(* Logix 5000 project; controller PLC_MCC1300_75F1 vendor 1 type 14 code 166 rev 32.11; software revision 32.04; part 66 of 83 *)
(* tags used below, declared in another part *)
   CM_ConveyorStackerToLine_JS1_Sync : CM_ConveyorStackerToLine;
   GP_AccessArea_M316S_STC : GP_AccessArea_STC;
   GP_ScadaPlate : GP_ScadaPlate;
   Gp_SpaceConvUtilities_V1 : GP_SpaceConvUtilities_V1;
   M310B : MAC_Conveyor;
   M312 : MAC_Conveyor_Single;
   M312_Data : UDT_Convoy_SL;
   M315A_SpaceConv_Utilities : SpaceConv_Utilities;
   M316 : MAC_Conveyor;
   M316_ALM : MAC_Conveyor_ALM;
   M316_Data : UDT_Convoy_SL;
   M316_HMR : MAC_Conveyor_HMR;
   M316_HMW : MAC_Conveyor_HMW;
   M316_M1_DR : AXIS_CIP_DRIVE;
   M316_SpaceConv_Utilities : SpaceConv_Utilities;
   M316_TON_Synchro_timeout : TIMER;
   M316_xSendCulletReqActive : BOOL;
   M316_xSensorTimeout : BOOL;
   M316A : MAC_Rotator;
   M316A_ALM : MAC_Rotator_ALM;
   M316A_Data : UDT_Convoy_SL;
   M316A_M1_DR_IN_MAM : MOTION_INSTRUCTION;
   M316A_TmON1 : TIMER;
   M316M317_OffsetBaricentre_cmm : DINT;
   M317 : MAC_Conveyor_Single;
   M317_ALM : MAC_Conveyor_ALM;
   M317_Data : UDT_Convoy_SL;
   M317_M2_DR_OUT_MAM : MOTION_INSTRUCTION;
   M317_M3_DR_OUT_MAM : MOTION_INSTRUCTION;
   M317_SpaceConv_Utilities : SpaceConv_Utilities;
   O : INT[128];
   TMP_d : DINT;
   TMP_SendToCullet : BOOL;
   TMP_xConveyorOfStartCleaning : BOOL;
   TMP_xEnableZoneCleaning : BOOL;
   TMP_xLiteThisDestPresent : BOOL;
   xAlwaysOFF : BOOL;
   xAlwaysON : BOOL;
   Z402 : MAC_Zone;
   Z402_HMI_rgtPlateScada_Internal : HMI_LiteData[5,2,7];
   Z402S_INPUT_xSafetyAreaPopup : BOOL;
   Z402S_INPUT_xSafetyAreaRotator : BOOL;
(* MainProgram, continued *)

   // Phase in progress
   48: NEQ(M316.PH_x,0)OTE(M316.ST_xPhasesInProgress);
   // #####_CLEANING_#####
   49: NOP();
   // Cleaning Reset
   50: XIC(M316.ST_xCleaningAccepted)[XIC(Z402.ST_xCleaningAccepted) ,XIO(TMP_xConveyorOfStartCleaning) ][XIC(M316.ST_xIdPlatePresence) OTL(TMP_SendToCullet) FLL(0,M316_Data,1) FLL(0,M316A_Data,1) ,MOV(0,M316A.PH_x) MOV(0,M316.PH_x) OTU(M316.ST_xPlatePresence) ];
   // Redestination lites
   // -
   // -
   51: [XIO(M316.ST_xPhasesInProgress) XIC(M312.ST_xAux1) ,XIC(M316_xSendCulletReqActive) [XIC(xAlwaysOFF) XIC(M316.PH_x.0) ,XIC(xAlwaysOFF) XIC(M316.PH_x.1) ,XIO(M316.ST_xPhasesInProgress) ] ]XIC(TMP_xLiteThisDestPresent)OTL(TMP_SendToCullet);
   // Initial condition OK
   52: XIC(Z402.ST_xConditionOkPhaseAdvancement)XIC(M316.ST_xOutputEnable)XIO(M316_HMW.xEnableDisableManualCommand)XIO(M316.ST_xReqCleaning)XIO(M316.ST_xCleaningAccepted)XIO(M316.ST_xStopNextCycleFault)XIO(M316.ST_xVirtualDoorEnabled)XIO(M316.PH_x.0)[XIO(M316.ST_xPhasesInProgress) XIO(M316.ST_xPlatePresence) XIO(M316.ST_xIdPlatePresence) XIC(M316A.INPUT_xLowPosition) ,XIC(M316.ST_xCycleLoadUnload) XIC(M316.PH_x.8) XIC(M316.OUTPUT_xRun_M1) GRT(M316_SpaceConv_Utilities.O_dTailPosition_cmm,M316_SpaceConv_Utilities.O_dPresetLoadUnload_cmm) GRT(M316_SpaceConv_Utilities.O_dTailPosition_cmm,380000) XIO(M316.ST_xIdPlatePresence) XIO(M312.INPUT_xSyncroPhotocell_1) ]XIO(CM_ConveyorStackerToLine_JS1_Sync.xRequestReturnInLine)XIO(GP_AccessArea_M316S_STC.ST_xAccessRequest)XIO(GP_AccessArea_M316S_STC.ST_xAccessAccepted)OTE(M316.ST_xInitialConditionOK);
   // #### Plate reentry ####
   53: NOP();
   // Initial condition reentry
   54: XIC(Z402.ST_xConditionOkPhaseAdvancement)XIC(M316.ST_xOutputEnable)XIO(M316_HMW.xEnableDisableManualCommand)XIO(M316.ST_xReqCleaning)XIO(M316.ST_xCleaningAccepted)XIO(M316.ST_xStopNextCycleFault)XIO(M312.ST_xVirtualDoorEnabled)XIO(M316.ST_xPhasesInProgress)XIO(M316.ST_xPlatePresence)XIO(M316.ST_xIdPlatePresence)XIC(M316A.INPUT_xLowPosition)XIO(GP_AccessArea_M316S_STC.ST_xAccessRequest)XIO(GP_AccessArea_M316S_STC.ST_xAccessAccepted)XIC(Z402S_INPUT_xSafetyAreaPopup)OTE(M316.ST_xInitialConditionOK_BW);
   // Phase of load reentry (backward)
   55: XIC(M312.OS_xUnload_BW)[OTL(M316.PH_x.22) ,OTU(M316_SpaceConv_Utilities.O_xPlateSynchronized) ,OTU(M316.ST_xDisableLoadUnloadOnStop) ,OTE(M316.OS_xLoad_BW) ,NEQ(M312_Data.rgtCap[0].rgtLite[0].dID,0) COP(M312_Data,M316_Data,1) FLL(0,M316_Data.rgtCap[0].rgtLite[1],1) ADD(M316_Data.rgtCap[0].rgtLite[0].dBarycenter_cmm,M316M317_OffsetBaricentre_cmm,M316_Data.rgtCap[0].rgtLite[0].dBarycenter_cmm) GP_SpaceConvUtilities_V1(Gp_SpaceConvUtilities_V1,M316_SpaceConv_Utilities,M315A_SpaceConv_Utilities,M317_SpaceConv_Utilities,15) ,FLL(0,M312_Data,1) ];
   // End load reentry (from M405) NEGATIVE
   56: XIC(M316.PH_x.22)[[GRT(M316_SpaceConv_Utilities.O_dHeadPosition_cmm,M316.AUX_dPresetStopLoad_cmm) XIO(M312.INPUT_xSyncroPhotocell_1) ,GRT(M316_SpaceConv_Utilities.O_dHeadPosition_cmm,450000) ] ,CPT(TMP_d,M316_SpaceConv_Utilities.CONST_dConveyorLength_cmm/2 + M316_Data.dLength_cmm / 2) GRT(M316_SpaceConv_Utilities.O_dHeadPosition_cmm,TMP_d) XIO(M312.INPUT_xSyncroPhotocell_1) ][OTE(M316.PH_x.23) ,OTU(M316.PH_x.22) ,OTL(M316.ST_xPlatePresence) ];
   // Phase of unload reentry (to M310B) NEGATIVE
   57: XIC(Z402.ST_xConditionOkPhaseAdvancement)XIC(M316.ST_xPlatePresence)XIC(M316.ST_xIdPlatePresence)XIO(TMP_xLiteThisDestPresent)XIC(M316.ST_xOutputEnable)XIO(M316.ST_xWaitMachineStop)XIO(M316.ST_xPhasesInProgress)[XIC(M310B.ST_xInitialConditionOK_BW) XIO(M316.ST_xVirtualDoorEnabled) [XIC(M316.ST_xAxleReadyToMoveDelayed) ,XIC(xAlwaysON) ] [XIC(M316.ST_xPlatePresence) XIC(M316.ST_xIdPlatePresence) OTE(M316.OS_xUnload_BW) ,OTL(M316.PH_x.24) ,XIC(M316.ST_xPlatePresence) XIC(M316.ST_xIdPlatePresence) MOV(M316_Data.dLength_cmm,M316_SpaceConv_Utilities.CONF_MD4_MD6_dLength_cmm) GP_SpaceConvUtilities_V1(Gp_SpaceConvUtilities_V1,M316_SpaceConv_Utilities,M315A_SpaceConv_Utilities,M317_SpaceConv_Utilities,16) ] ,OTE(M316.ST_xAux1) ];
   // Phase of end unload (to M310B) NEGATIVE
   58: XIC(M316.PH_x.24)[[GEQ(M316_SpaceConv_Utilities.O_dTailPosition_cmm,M316.AUX_dPresetStopUnload_cmm) ,LEQ(M316_SpaceConv_Utilities.O_dTailPosition_cmm,0) GEQ(M316_SpaceConv_Utilities.O_dTailPosition_cmm,M316.AUX_dPresetStopUnload_cmm) ] ,XIO(M316_SpaceConv_Utilities.ST_xFeedbackRotation) GEQ(M316_SpaceConv_Utilities.O_dTailPosition_cmm,M316_SpaceConv_Utilities.CONST_dConveyorLength_cmm) ,XIO(xAlwaysOFF) XIC(M310B.PH_x.29) ][OTE(M316.PH_x.25) ,OTU(M316.PH_x.24) ,OTU(M316.ST_xPlatePresence) ];
   // #####_HMI_STATUSES_#####
   59: NOP();
   // PhotocelPresence {x|x|x|x|O}
   60: XIC(M316.INPUT_xSyncroPhotocell_1)OTE(M316_HMR.xSensorPresence1);
   // PhotocelPresence {x|x|x|x|O}
   61: XIC(M316.INPUT_xSyncroPhotocell_2)OTE(M316_HMR.xSensorPresence2);
   // Manual Mode Enable {x|x|x|x|O}
   62: XIC(M316.ST_xManualMode)OTE(M316_HMR.xManualCommandEnabled);
   // Command forward M1
   63: XIC(M316.ST_xManualMode)XIC(M316_HMW.rgxMan.0)XIC(M316.OUTPUT_xRun_M1)OTE(M316_HMR.rgxMan.0);
   // Command backward M1
   64: XIC(M316.ST_xManualMode)XIC(M316_HMW.rgxMan.1)XIC(M316.OUTPUT_xReverse_M1)OTE(M316_HMR.rgxMan.1);
   // Command forward M2
   65: XIC(M316.ST_xManualMode)XIC(M316_HMW.rgxMan.2)XIC(M316.OUTPUT_xRun_M2)OTE(M316_HMR.rgxMan.2);
   // Command backward M2
   66: XIC(M316.ST_xManualMode)XIC(M316_HMW.rgxMan.3)XIC(M316.OUTPUT_xReverse_M2)OTE(M316_HMR.rgxMan.3);
   // Cleaning Enabled {x|x|x|x|O}
   67: XIC(M316.ST_xCleaningAccepted)[XIC(Z402.ST_xCleaningAccepted) ,XIO(TMP_xEnableZoneCleaning) ]OTE(M316_HMR.xCleaningEnabled);
   // Virtual door Enabled {x|x|x|x|O}
   68: XIC(M316.ST_xVirtualDoorEnabled)OTE(M316_HMR.xVirtualDoorEnabled);
   // Id plate presence
   69: XIC(M316.ST_xIdPlatePresence)OTE(M316_HMR.xIdPlatePresence);
   // Machine state M1
   70: XIC(xAlwaysON)[MOV(1,M316_HMR.dState1) ,XIC(M316.OUTPUT_xRun_M1) MOV(3,M316_HMR.dState1) ,XIC(M316.OUTPUT_xReverse_M1) MOV(4,M316_HMR.dState1) ,XIC(M316.ST_xMachineAlarm) MOV(7,M316_HMR.dState1) ];
   // Machine state M2
   71: XIC(xAlwaysON)[MOV(1,M316_HMR.dState2) ,XIC(M316.OUTPUT_xRun_M2) MOV(3,M316_HMR.dState2) ,XIC(M316.OUTPUT_xReverse_M2) MOV(4,M316_HMR.dState2) ,XIC(M316.ST_xMachineAlarm) MOV(7,M316_HMR.dState2) ];
   72: XIC(M316.INPUT_xSyncroPhotocell_1)XIO(M316.ST_xIdPlatePresence)XIO(M316.ST_xPlatePresence)[TON(M316_TON_Synchro_timeout,?,?) ,[XIC(M316_TON_Synchro_timeout.DN) ,XIC(M316_xSensorTimeout) ] XIC(M316.INPUT_xSyncroPhotocell_1) OTE(M316_xSensorTimeout) ];
   // State Sensor
   73: XIC(xAlwaysON)[MOV(1,M316_HMR.dStateSensor1) ,[XIC(M316_ALM.rgxWarning[0].0) ,XIC(M316_xSensorTimeout) ] MOV(7,M316_HMR.dStateSensor1) ];
   // State Sensor
   74: XIC(xAlwaysON)[MOV(1,M316_HMR.dStateSensor2) ,XIC(M316_ALM.rgxWarning[0].1) MOV(7,M316_HMR.dStateSensor2) ];
   // State Sensor
   75: XIC(xAlwaysON)[MOV(1,M316_HMR.dStateSensor3) ,XIC(M316_ALM.rgxWarning[0].0) MOV(7,M316_HMR.dStateSensor3) ];
   // State Sensor
   76: XIC(xAlwaysON)[MOV(1,M316_HMR.dStateSensor4) ,XIC(M316_ALM.rgxWarning[0].1) MOV(7,M316_HMR.dStateSensor4) ];
   // Motor error code
   77: MOV(M316_M1_DR.AxisFault,M316_HMR.dErrorCode1);
   78: XIC(M316.ST_xIdPlatePresence)GP_ScadaPlate(GP_ScadaPlate,M316_Data,2,M316_SpaceConv_Utilities.O_dHeadPosition_cmm,M316_SpaceConv_Utilities.CONST_dConveyorWidth_cmm,M316_SpaceConv_Utilities.CONST_dConveyorLength_cmm,M316_SpaceConv_Utilities.ST_xLastModLoadBkw,M316_SpaceConv_Utilities.ST_xLastModUnloadBkw,1,0,Z402_HMI_rgtPlateScada_Internal);
END_ROUTINE

ROUTINE M316A_Rotator_Alarm   (* ladder *)
   // Reset Alarm
   0: XIC(Z402.tmON_ResetAlarm.DN)FLL(0,M316A_ALM,1);
   1: XIC(Z402.ST_xEnableControlError)XIC(M316A.INPUT_xProtectionMotorRotation)XIC(M316A.INPUT_xProtectionMotorLifting)OTE(M316A.ST_xEnableControlError);
   2: XIC(Z402.ST_xEnableControlError)XIO(M316A.INPUT_xProtectionMotorRotation)OTL(M316A_ALM.rgxStoppingFault_M[0].0);
   3: XIC(M316A.ST_xEnableControlError)XIC(M316A.INPUT_xDriveError)OTL(M316A_ALM.rgxStoppingFault_M[0].1);
   4: XIC(M316A.ST_xEnableControlError)XIO(M316A.INPUT_xDriveError)[XIC(M316A.OUTPUT_xRun) ,XIC(M316A.OUTPUT_xReverse) ][XIO(M316A_M1_DR_IN_MAM.EN) ,XIC(M316A_M1_DR_IN_MAM.EN) XIO(M316A_M1_DR_IN_MAM.PC) ]XIO(M316A.INPUT_xDriveFeedback)[XIO(M316A.tmON_FeedbackTimeOutRotation.DN) TON(M316A.tmON_FeedbackTimeOutRotation,?,?) ,XIC(M316A.tmON_FeedbackTimeOutRotation.DN) OTL(M316A_ALM.rgxStoppingFault_M[0].2) ];
   5: XIC(M316A.ST_xEnableControlError)[XIC(M316A_M1_DR_IN_MAM.IP) TON(M316A.tmON_RotatePosError,?,?) ,[XIC(M316A.tmON_RotatePosError.DN) ,XIO(M316A.OUTPUT_xRun) XIO(M316A.OUTPUT_xReverse) XIO(M316A.ST_xFeedbackRotation) XIO(M316A.INPUT_xConditionToDescent) ] OTL(M316A_ALM.rgxStoppingFault_M[0].3) ];
   6: XIC(Z402.ST_xEnableControlError)XIO(M316A.INPUT_xLocalSafetySwitchRotation)XIC(xAlwaysOFF)OTL(M316A_ALM.rgxStoppingFault_M[0].4);
   7: XIC(Z402.ST_xEnableControlError)XIO(M316A.INPUT_xBrakingResistor)XIC(xAlwaysOFF)OTL(M316A_ALM.rgxStoppingFault_M[0].5);
   8: XIC(Z402.ST_xEnableControlError)XIC(M316A.INPUT_xMotorThermalProbe)XIC(xAlwaysOFF)OTL(M316A_ALM.rgxStoppingFault_M[0].6);
   9: XIC(Z402.ST_xEnableControlError)XIO(M316A.INPUT_xProtectionMotorLifting)OTL(M316A_ALM.rgxStoppingFault_M[0].8);
   10: XIC(Z402.ST_xEnableControlError)XIC(Z402S_INPUT_xSafetyAreaRotator)[XIC(M316A.INPUT_xDriveInhibit) ,XIC(M316A.OUTPUT_xDriveEnable) XIO(M316A.INPUT_xDriveReady) ][XIO(M316A_TmON1.DN) TON(M316A_TmON1,?,?) ,XIC(M316A_TmON1.DN) OTL(M316A_ALM.rgxStoppingFault_M[0].20) ];
   11: XIC(M316A.ST_xEnableControlError)[[XIC(M316A.OUTPUT_xRise) ,XIC(M316A.OUTPUT_xDescent) ] XIO(M316A.INPUT_xFeedbackLifting) ,XIO(M316A.OUTPUT_xRise) XIO(M316A.OUTPUT_xDescent) XIC(M316A.INPUT_xFeedbackLifting) ][XIO(M316A.tmON_FeedbackTimeOutLifting.DN) TON(M316A.tmON_FeedbackTimeOutLifting,?,?) ,XIC(M316A.tmON_FeedbackTimeOutLifting.DN) OTL(M316A_ALM.rgxStoppingFault_M[0].9) ];
   12: XIC(M316A.ST_xEnableControlError)[[XIC(M316A.OUTPUT_xRise) XIO(M316A.INPUT_xHighPosition) ,XIC(M316A.OUTPUT_xDescent) XIO(M316A.INPUT_xLowPosition) ,XIO(M316A.INPUT_xHighPosition) XIO(M316A.INPUT_xLowPosition) ] XIO(M316A.tmON_FramePosError.DN) TON(M316A.tmON_FramePosError,?,?) ,[XIC(M316A.tmON_FramePosError.DN) ,XIC(M316A.INPUT_xHighPosition) XIC(M316A.INPUT_xLowPosition) ] OTL(M316A_ALM.rgxStoppingFault_M[0].11) ];
   13: XIC(Z402.ST_xEnableControlError)XIO(M316A.INPUT_xLocalSafetySwitchLifting)XIC(xAlwaysOFF)OTL(M316A_ALM.rgxStoppingFault_M[0].12);
   // #####_CUMULATIVE ALARM_#####
   14: NOP();
   15: [NEQ(M316A_ALM.rgxStoppingFault[0],0) ,NEQ(M316A_ALM.rgxStoppingFault_M[0],0) ]OTE(M316A.ST_xStopMachineFault);
   16: [NEQ(M316A_ALM.rgxFault[0],0) ,NEQ(M316A_ALM.rgxFault_M[0],0) ]OTE(M316A.ST_xStopNextCycleFault);
END_ROUTINE

ROUTINE M317_Alarm   (* ladder *)
   // Reset Alarm
   0: XIC(Z402.tmON_ResetAlarm.DN)FLL(0,M317_ALM,1);
   // M1
   // -
   // -
   1: NOP();
   2: XIC(Z402.ST_xEnableControlError)XIC(xAlwaysOFF)XIO(M317.INPUT_xProtectionMotor_M1)OTL(M317_ALM.rgxStoppingFault_M[0].0);
   3: XIC(Z402.ST_xEnableControlError)XIC(M317.INPUT_xDriveError_M1)OTL(M317_ALM.rgxStoppingFault_M[0].1);
   4: XIC(Z402.ST_xEnableControlError)XIO(M317.INPUT_xDriveError_M1)[XIC(M317.OUTPUT_xRun_M1) ,XIC(M317.OUTPUT_xReverse_M1) ,XIC(M317.OUTPUT_xPositioning_M1) ]XIO(M317.INPUT_xDriveFeedback_M1)[XIO(M317.tmON_FeedbackTimeOut_M1.DN) TON(M317.tmON_FeedbackTimeOut_M1,?,?) ,XIC(M317.tmON_FeedbackTimeOut_M1.DN) OTL(M317_ALM.rgxStoppingFault_M[0].2) ];
   5: XIC(Z402.ST_xEnableControlError)XIC(xAlwaysOFF)XIO(M317.INPUT_xLocalSafetySwitch_M1)OTL(M317_ALM.rgxStoppingFault_M[0].3);
   6: XIC(Z402.ST_xEnableControlError)XIO(M317.INPUT_xMotorThermalProbe_M1)OTL(M317_ALM.rgxStoppingFault_M[0].4);
   7: XIC(Z402.ST_xEnableControlError)XIC(xAlwaysOFF)XIO(M317.INPUT_xBrakingResistor_M1)OTL(M317_ALM.rgxStoppingFault_M[0].5);
   8: XIC(Z402.ST_xEnableControlError)[XIC(M317.INPUT_xDriveInhibit_M1) ,XIC(M317.OUTPUT_xDriveEnable_M1) XIO(M317.INPUT_xDriveReady_M1) ][XIO(M317.TmON[11].DN) TON(M317.TmON[11],?,?) ,XIC(M317.TmON[11].DN) OTL(M317_ALM.rgxStoppingFault_M[0].6) ];
   9: XIC(xAlwaysOFF)XIC(M317.ST_xEnableControlError)XIC(M317.PH_x.7)NEQ(M317_SpaceConv_Utilities.CONST_dSyncMode,0)[XIO(M317.ST_xPlateSynchronized) OTL(M317_ALM.rgxWarning[0].0) ,XIC(M317.ST_xPlateSynchronized) OTU(M317_ALM.rgxWarning[0].0) ];
   10: XIC(M317.ST_xEnableControlError)XIC(M317_Data.tFlag.tConveyor.xReqStop)XIC(M317.PH_x.0)GRT(M317_SpaceConv_Utilities.O_dHeadPosition_cmm,M317_SpaceConv_Utilities.CONST_dConveyorLength_cmm)[OTL(M317_ALM.rgxWarning[0].1) ,OTL(M317.ST_xPhaseError) ];
   // M2
   // -
   // -
   11: NOP();
   12: XIC(Z402.ST_xEnableControlError)XIC(xAlwaysOFF)XIO(M317.INPUT_xProtectionMotor_M2)OTL(M317_ALM.rgxStoppingFault_M[0].8);
   13: XIC(Z402.ST_xEnableControlError)XIC(M317.INPUT_xDriveError_M2)OTL(M317_ALM.rgxStoppingFault_M[0].9);
   14: XIC(Z402.ST_xEnableControlError)XIO(M317.INPUT_xDriveError_M2)[XIC(M317.OUTPUT_xRun_M2) ,XIC(M317.OUTPUT_xReverse_M2) ,XIC(M317.OUTPUT_xPositioning_M2) XIO(M317_M2_DR_OUT_MAM.DN) ]XIO(M317.INPUT_xDriveFeedback_M2)[XIO(M317.tmON_FeedbackTimeOut_M2.DN) TON(M317.tmON_FeedbackTimeOut_M2,?,?) ,XIC(M317.tmON_FeedbackTimeOut_M2.DN) OTL(M317_ALM.rgxStoppingFault_M[0].10) ];
   15: XIC(Z402.ST_xEnableControlError)XIC(xAlwaysOFF)XIO(M317.INPUT_xLocalSafetySwitch_M2)OTL(M317_ALM.rgxStoppingFault_M[0].11);
   16: XIC(Z402.ST_xEnableControlError)XIO(M317.INPUT_xMotorThermalProbe_M2)OTL(M317_ALM.rgxStoppingFault_M[0].12);
   17: XIC(Z402.ST_xEnableControlError)XIC(xAlwaysOFF)XIO(M317.INPUT_xBrakingResistor_M2)OTL(M317_ALM.rgxStoppingFault_M[0].13);
   18: XIC(Z402.ST_xEnableControlError)[XIC(M317.INPUT_xDriveInhibit_M2) ,XIC(M317.OUTPUT_xDriveEnable_M2) XIO(M317.INPUT_xDriveReady_M2) ][XIO(M317.TmON[12].DN) TON(M317.TmON[12],?,?) ,XIC(M317.TmON[12].DN) OTL(M317_ALM.rgxStoppingFault_M[0].14) ];
   19: XIC(Z402.ST_xEnableControlError)[XIC(M317.ST_xOutputEnable) [XIC(M317.PH_x.24) ,XIC(M317.PH_x.26) ] XIO(M317.tmON_AuxFunction4.DN) TON(M317.tmON_AuxFunction4,?,?) ,XIC(M317.tmON_AuxFunction4.DN) [OTL(M317_ALM.rgxWarning[0].11) ,OTL(M317.ST_xPhaseError) ] ];
   // M3
   // -
   // -
   20: NOP();
   21: XIC(Z402.ST_xEnableControlError)XIC(xAlwaysOFF)XIO(M317.INPUT_xProtectionMotor_M3)OTL(M317_ALM.rgxStoppingFault_M[0].16);
   22: XIC(Z402.ST_xEnableControlError)XIC(M317.INPUT_xDriveError_M3)OTL(M317_ALM.rgxStoppingFault_M[0].17);
   23: XIC(Z402.ST_xEnableControlError)XIO(M317.INPUT_xDriveError_M3)[XIC(M317.OUTPUT_xRun_M3) ,XIC(M317.OUTPUT_xReverse_M3) ,XIC(M317.OUTPUT_xPositioning_M3) XIO(M317_M3_DR_OUT_MAM.DN) ]XIO(M317.INPUT_xDriveFeedback_M3)[XIO(M317.tmON_FeedbackTimeOut_M3.DN) TON(M317.tmON_FeedbackTimeOut_M3,?,?) ,XIC(M317.tmON_FeedbackTimeOut_M3.DN) OTL(M317_ALM.rgxStoppingFault_M[0].18) ];
   24: XIC(Z402.ST_xEnableControlError)XIC(xAlwaysOFF)XIO(M317.INPUT_xLocalSafetySwitch_M3)OTL(M317_ALM.rgxStoppingFault_M[0].19);
   25: XIC(Z402.ST_xEnableControlError)XIO(M317.INPUT_xMotorThermalProbe_M3)OTL(M317_ALM.rgxStoppingFault_M[0].20);
   26: XIC(Z402.ST_xEnableControlError)XIC(xAlwaysOFF)XIO(M317.INPUT_xBrakingResistor_M3)OTL(M317_ALM.rgxStoppingFault_M[0].21);
   27: XIC(Z402.ST_xEnableControlError)XIC(Z402S_INPUT_xSafetyAreaRotator)[XIC(M317.INPUT_xDriveInhibit_M3) ,XIC(M317.OUTPUT_xDriveEnable_M3) XIO(M317.INPUT_xDriveReady_M3) ][XIO(M317.TmON[13].DN) TON(M317.TmON[13],?,?) ,XIC(M317.TmON[13].DN) OTL(M317_ALM.rgxStoppingFault_M[0].21) ];
   // M4
   // -
   // -
   28: NOP();
   29: XIC(Z402.ST_xEnableControlError)XIC(xAlwaysOFF)XIO(M317.INPUT_xProtectionMotor_M4)OTL(M317_ALM.rgxStoppingFault_M[0].24);
   30: XIC(Z402.ST_xEnableControlError)XIC(M317.INPUT_xDriveError_M4)OTL(M317_ALM.rgxStoppingFault_M[0].25);
   31: XIC(Z402.ST_xEnableControlError)XIO(M317.INPUT_xMotorThermalProbe_M4)OTL(M317_ALM.rgxStoppingFault_M[0].28);
